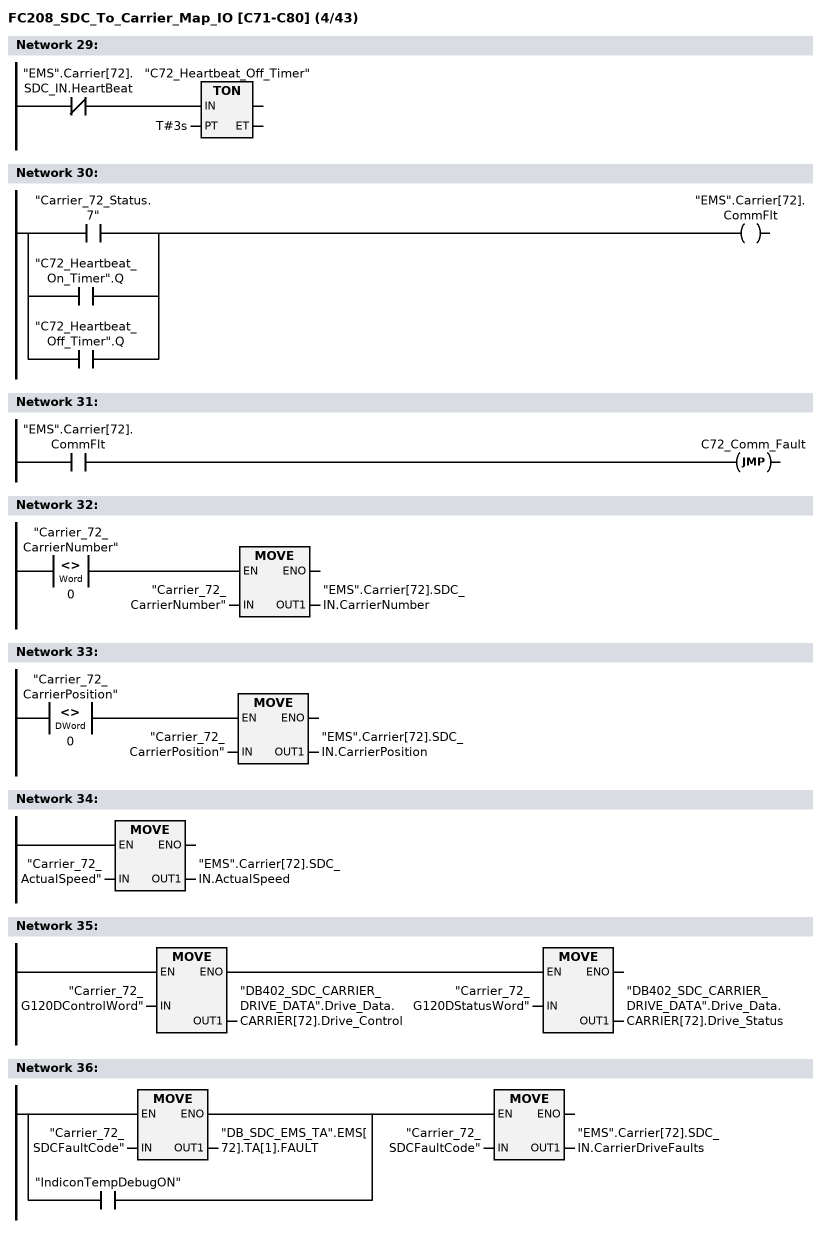
   "C72_Heartbeat_Off_Timer".TON(IN := NOT "EMS".Carrier[72].SDC_IN.HeartBeat, PT := T#3s);
END_REGION

REGION Network 30
   RUNG wire#powerrail
      Contact( "Carrier_72_Status.7" )
      wire#w1
      Coil( "EMS".Carrier[72].CommFlt )
   END_RUNG
   RUNG wire#powerrail
      Contact( "C72_Heartbeat_On_Timer".Q )
   END_RUNG wire#w1
   RUNG wire#powerrail
      Contact( "C72_Heartbeat_Off_Timer".Q )
   END_RUNG wire#w1
   // the same network as SCL:
   "EMS".Carrier[72].CommFlt := "Carrier_72_Status.7" OR "C72_Heartbeat_On_Timer".Q OR "C72_Heartbeat_Off_Timer".Q;
END_REGION

REGION Network 31
   RUNG wire#powerrail
      Contact( "EMS".Carrier[72].CommFlt )
      JumpCoil( C72_Comm_Fault )
   END_RUNG
   // the same network as SCL:
   IF "EMS".Carrier[72].CommFlt THEN GOTO C72_Comm_Fault; END_IF;
END_REGION

REGION Network 32
   RUNG wire#powerrail
      { S7_Templates := "SrcType := Word" } NE_Contact(in1 := "Carrier_72_CarrierNumber", in2 := 0)
      Move(in := "Carrier_72_CarrierNumber", out1 => "EMS".Carrier[72].SDC_IN.CarrierNumber)
   END_RUNG
   // the same network as SCL:
   IF "Carrier_72_CarrierNumber" <> 0 THEN
       "EMS".Carrier[72].SDC_IN.CarrierNumber := "Carrier_72_CarrierNumber";
   END_IF;
END_REGION

REGION Network 33
   RUNG wire#powerrail
      { S7_Templates := "SrcType := DWord" } NE_Contact(in1 := "Carrier_72_CarrierPosition", in2 := 0)
      Move(in := "Carrier_72_CarrierPosition", out1 => "EMS".Carrier[72].SDC_IN.CarrierPosition)
   END_RUNG
   // the same network as SCL:
   IF "Carrier_72_CarrierPosition" <> 0 THEN
       "EMS".Carrier[72].SDC_IN.CarrierPosition := "Carrier_72_CarrierPosition";
   END_IF;
END_REGION

REGION Network 34
   RUNG wire#powerrail
      Move(in := "Carrier_72_ActualSpeed", out1 => "EMS".Carrier[72].SDC_IN.ActualSpeed)
   END_RUNG
   // the same network as SCL:
   "EMS".Carrier[72].SDC_IN.ActualSpeed := "Carrier_72_ActualSpeed";
END_REGION

REGION Network 35
   RUNG wire#powerrail
      Move(in := "Carrier_72_G120DControlWord", out1 => "DB402_SDC_CARRIER_DRIVE_DATA".Drive_Data.CARRIER[72].Drive_Control)
      Move(in := "Carrier_72_G120DStatusWord", out1 => "DB402_SDC_CARRIER_DRIVE_DATA".Drive_Data.CARRIER[72].Drive_Status)
   END_RUNG
   // the same network as SCL:
   "DB402_SDC_CARRIER_DRIVE_DATA".Drive_Data.CARRIER[72].Drive_Control := "Carrier_72_G120DControlWord";
   "DB402_SDC_CARRIER_DRIVE_DATA".Drive_Data.CARRIER[72].Drive_Status := "Carrier_72_G120DStatusWord";
END_REGION

REGION Network 36
   RUNG wire#powerrail
      Move(in := "Carrier_72_SDCFaultCode", out1 => "DB_SDC_EMS_TA".EMS[72].TA[1].FAULT)
      wire#w1
      Move(in := "Carrier_72_SDCFaultCode", out1 => "EMS".Carrier[72].SDC_IN.CarrierDriveFaults)
   END_RUNG
   RUNG wire#powerrail
      Contact( "IndiconTempDebugON" )
   END_RUNG wire#w1
   // the same network as SCL:
   "DB_SDC_EMS_TA".EMS[72].TA[1].FAULT := "Carrier_72_SDCFaultCode";
   IF TRUE OR "IndiconTempDebugON" THEN
       "EMS".Carrier[72].SDC_IN.CarrierDriveFaults := "Carrier_72_SDCFaultCode";
   END_IF;
END_REGION

REGION Network 37
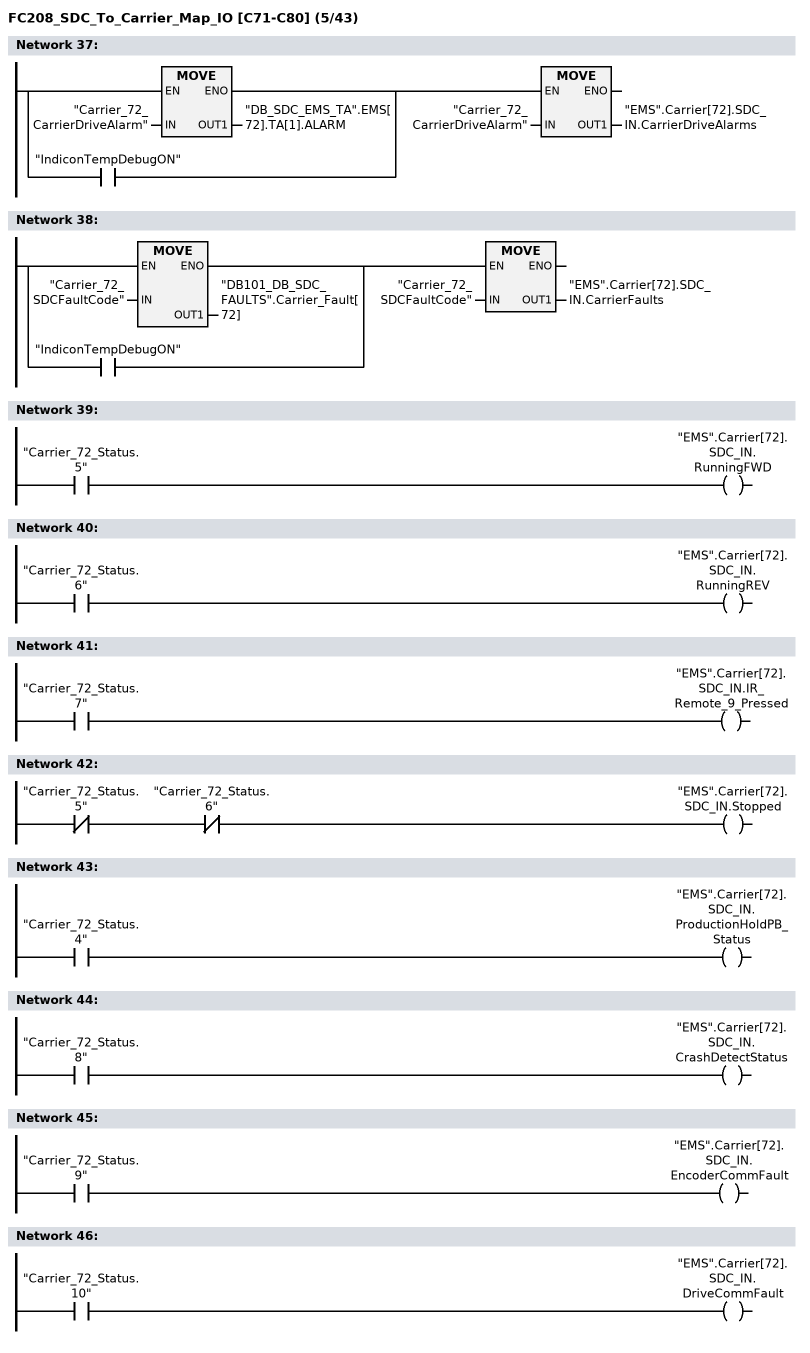
   RUNG wire#powerrail
      Move(in := "Carrier_72_CarrierDriveAlarm", out1 => "DB_SDC_EMS_TA".EMS[72].TA[1].ALARM)
      wire#w1
      Move(in := "Carrier_72_CarrierDriveAlarm", out1 => "EMS".Carrier[72].SDC_IN.CarrierDriveAlarms)
   END_RUNG
   RUNG wire#powerrail
      Contact( "IndiconTempDebugON" )
   END_RUNG wire#w1
   // the same network as SCL:
   "DB_SDC_EMS_TA".EMS[72].TA[1].ALARM := "Carrier_72_CarrierDriveAlarm";
   IF TRUE OR "IndiconTempDebugON" THEN
       "EMS".Carrier[72].SDC_IN.CarrierDriveAlarms := "Carrier_72_CarrierDriveAlarm";
   END_IF;
END_REGION

REGION Network 38
   RUNG wire#powerrail
      Move(in := "Carrier_72_SDCFaultCode", out1 => "DB101_DB_SDC_FAULTS".Carrier_Fault[72])
      wire#w1
      Move(in := "Carrier_72_SDCFaultCode", out1 => "EMS".Carrier[72].SDC_IN.CarrierFaults)
   END_RUNG
   RUNG wire#powerrail
      Contact( "IndiconTempDebugON" )
   END_RUNG wire#w1
   // the same network as SCL:
   "DB101_DB_SDC_FAULTS".Carrier_Fault[72] := "Carrier_72_SDCFaultCode";
   IF TRUE OR "IndiconTempDebugON" THEN
       "EMS".Carrier[72].SDC_IN.CarrierFaults := "Carrier_72_SDCFaultCode";
   END_IF;
END_REGION

REGION Network 39
   RUNG wire#powerrail
      Contact( "Carrier_72_Status.5" )
      Coil( "EMS".Carrier[72].SDC_IN.RunningFWD )
   END_RUNG
   // the same network as SCL:
   "EMS".Carrier[72].SDC_IN.RunningFWD := "Carrier_72_Status.5";
END_REGION

REGION Network 40
   RUNG wire#powerrail
      Contact( "Carrier_72_Status.6" )
      Coil( "EMS".Carrier[72].SDC_IN.RunningREV )
   END_RUNG
   // the same network as SCL:
   "EMS".Carrier[72].SDC_IN.RunningREV := "Carrier_72_Status.6";
END_REGION

REGION Network 41
   RUNG wire#powerrail
      Contact( "Carrier_72_Status.7" )
      Coil( "EMS".Carrier[72].SDC_IN.IR_Remote_9_Pressed )
   END_RUNG
   // the same network as SCL:
   "EMS".Carrier[72].SDC_IN.IR_Remote_9_Pressed := "Carrier_72_Status.7";
END_REGION

REGION Network 42
   RUNG wire#powerrail
      I_Contact( "Carrier_72_Status.5" )
      I_Contact( "Carrier_72_Status.6" )
      Coil( "EMS".Carrier[72].SDC_IN.Stopped )
   END_RUNG
   // the same network as SCL:
   "EMS".Carrier[72].SDC_IN.Stopped := NOT "Carrier_72_Status.5" AND NOT "Carrier_72_Status.6";
END_REGION

REGION Network 43
   RUNG wire#powerrail
      Contact( "Carrier_72_Status.4" )
      Coil( "EMS".Carrier[72].SDC_IN.ProductionHoldPB_Status )
   END_RUNG
   // the same network as SCL:
   "EMS".Carrier[72].SDC_IN.ProductionHoldPB_Status := "Carrier_72_Status.4";
END_REGION

REGION Network 44
   RUNG wire#powerrail
      Contact( "Carrier_72_Status.8" )
      Coil( "EMS".Carrier[72].SDC_IN.CrashDetectStatus )
   END_RUNG
   // the same network as SCL:
   "EMS".Carrier[72].SDC_IN.CrashDetectStatus := "Carrier_72_Status.8";
END_REGION

REGION Network 45
   RUNG wire#powerrail
      Contact( "Carrier_72_Status.9" )
      Coil( "EMS".Carrier[72].SDC_IN.EncoderCommFault )
   END_RUNG
   // the same network as SCL:
   "EMS".Carrier[72].SDC_IN.EncoderCommFault := "Carrier_72_Status.9";
END_REGION

REGION Network 46
   RUNG wire#powerrail
      Contact( "Carrier_72_Status.10" )
      Coil( "EMS".Carrier[72].SDC_IN.DriveCommFault )
   END_RUNG
   // the same network as SCL:
   "EMS".Carrier[72].SDC_IN.DriveCommFault := "Carrier_72_Status.10";
END_REGION

REGION Network 47
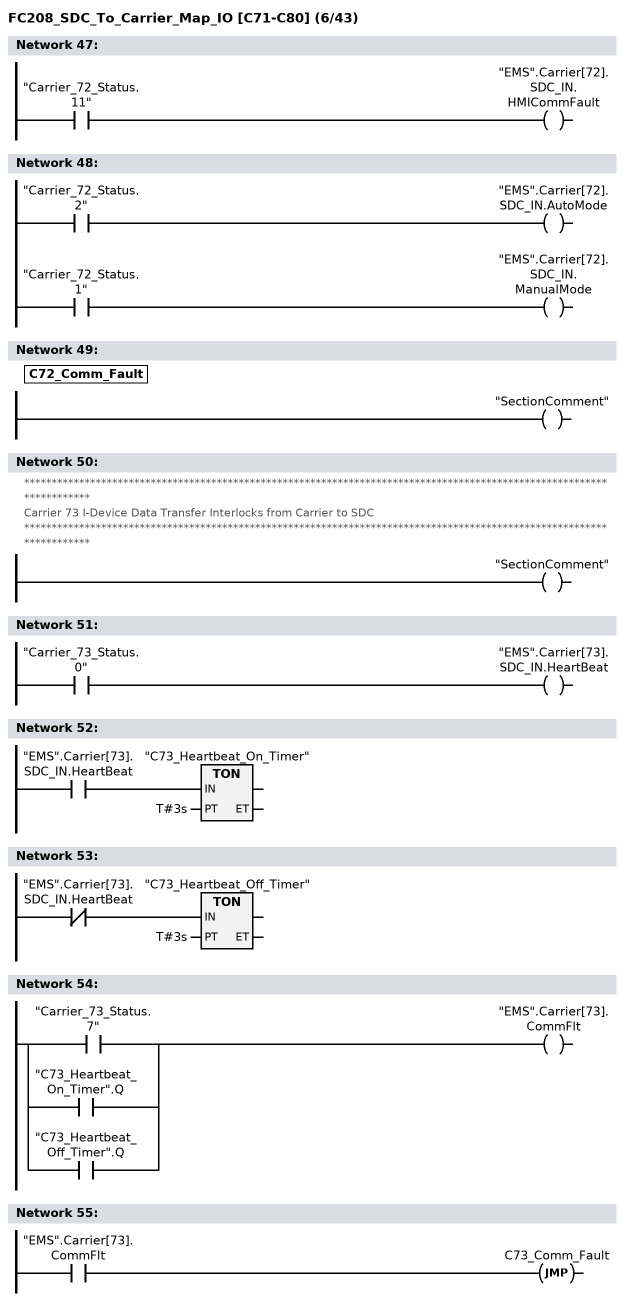
   RUNG wire#powerrail
      Contact( "Carrier_72_Status.11" )
      Coil( "EMS".Carrier[72].SDC_IN.HMICommFault )
   END_RUNG
   // the same network as SCL:
   "EMS".Carrier[72].SDC_IN.HMICommFault := "Carrier_72_Status.11";
END_REGION

REGION Network 48
   RUNG wire#powerrail
      Contact( "Carrier_72_Status.2" )
      Coil( "EMS".Carrier[72].SDC_IN.AutoMode )
   END_RUNG
   RUNG wire#powerrail
      Contact( "Carrier_72_Status.1" )
      Coil( "EMS".Carrier[72].SDC_IN.ManualMode )
   END_RUNG
   // the same network as SCL:
   "EMS".Carrier[72].SDC_IN.AutoMode := "Carrier_72_Status.2";
   "EMS".Carrier[72].SDC_IN.ManualMode := "Carrier_72_Status.1";
END_REGION

REGION Network 49
   Label( C72_Comm_Fault )
   RUNG wire#powerrail
      Coil( "SectionComment" )
   END_RUNG
   // the same network as SCL:
   C72_Comm_Fault:
   "SectionComment" := TRUE;
END_REGION

REGION Network 50
   // **********************************************************************************************************************
   // 
   // Carrier 73 I-Device Data Transfer Interlocks from Carrier to SDC
   // 
   // **********************************************************************************************************************
   RUNG wire#powerrail
      Coil( "SectionComment" )
   END_RUNG
   // the same network as SCL:
   "SectionComment" := TRUE;
END_REGION

REGION Network 51
   RUNG wire#powerrail
      Contact( "Carrier_73_Status.0" )
      Coil( "EMS".Carrier[73].SDC_IN.HeartBeat )
   END_RUNG
   // the same network as SCL:
   "EMS".Carrier[73].SDC_IN.HeartBeat := "Carrier_73_Status.0";
END_REGION

REGION Network 52
   "C73_Heartbeat_On_Timer".TON(IN := "EMS".Carrier[73].SDC_IN.HeartBeat, PT := T#3s);
END_REGION

REGION Network 53
   "C73_Heartbeat_Off_Timer".TON(IN := NOT "EMS".Carrier[73].SDC_IN.HeartBeat, PT := T#3s);
END_REGION

REGION Network 54
   RUNG wire#powerrail
      Contact( "Carrier_73_Status.7" )
      wire#w1
      Coil( "EMS".Carrier[73].CommFlt )
   END_RUNG
   RUNG wire#powerrail
      Contact( "C73_Heartbeat_On_Timer".Q )
   END_RUNG wire#w1
   RUNG wire#powerrail
      Contact( "C73_Heartbeat_Off_Timer".Q )
   END_RUNG wire#w1
   // the same network as SCL:
   "EMS".Carrier[73].CommFlt := "Carrier_73_Status.7" OR "C73_Heartbeat_On_Timer".Q OR "C73_Heartbeat_Off_Timer".Q;
END_REGION

REGION Network 55
   RUNG wire#powerrail
      Contact( "EMS".Carrier[73].CommFlt )
      JumpCoil( C73_Comm_Fault )
   END_RUNG
   // the same network as SCL:
   IF "EMS".Carrier[73].CommFlt THEN GOTO C73_Comm_Fault; END_IF;
END_REGION

REGION Network 56
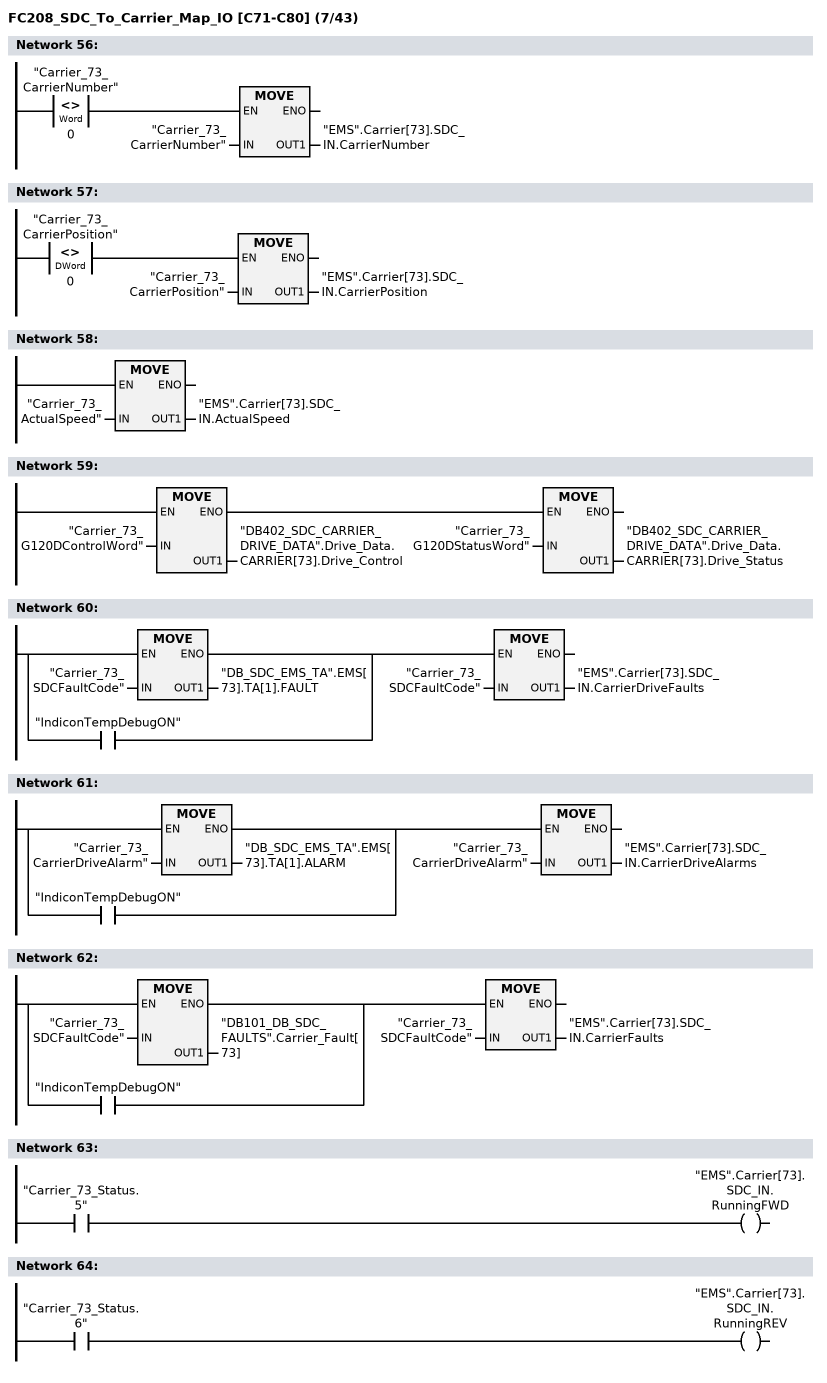
   RUNG wire#powerrail
      { S7_Templates := "SrcType := Word" } NE_Contact(in1 := "Carrier_73_CarrierNumber", in2 := 0)
      Move(in := "Carrier_73_CarrierNumber", out1 => "EMS".Carrier[73].SDC_IN.CarrierNumber)
   END_RUNG
   // the same network as SCL:
   IF "Carrier_73_CarrierNumber" <> 0 THEN
       "EMS".Carrier[73].SDC_IN.CarrierNumber := "Carrier_73_CarrierNumber";
   END_IF;
END_REGION

REGION Network 57
   RUNG wire#powerrail
      { S7_Templates := "SrcType := DWord" } NE_Contact(in1 := "Carrier_73_CarrierPosition", in2 := 0)
      Move(in := "Carrier_73_CarrierPosition", out1 => "EMS".Carrier[73].SDC_IN.CarrierPosition)
   END_RUNG
   // the same network as SCL:
   IF "Carrier_73_CarrierPosition" <> 0 THEN
       "EMS".Carrier[73].SDC_IN.CarrierPosition := "Carrier_73_CarrierPosition";
   END_IF;
END_REGION

REGION Network 58
   RUNG wire#powerrail
      Move(in := "Carrier_73_ActualSpeed", out1 => "EMS".Carrier[73].SDC_IN.ActualSpeed)
   END_RUNG
   // the same network as SCL:
   "EMS".Carrier[73].SDC_IN.ActualSpeed := "Carrier_73_ActualSpeed";
END_REGION

REGION Network 59
   RUNG wire#powerrail
      Move(in := "Carrier_73_G120DControlWord", out1 => "DB402_SDC_CARRIER_DRIVE_DATA".Drive_Data.CARRIER[73].Drive_Control)
      Move(in := "Carrier_73_G120DStatusWord", out1 => "DB402_SDC_CARRIER_DRIVE_DATA".Drive_Data.CARRIER[73].Drive_Status)
   END_RUNG
   // the same network as SCL:
   "DB402_SDC_CARRIER_DRIVE_DATA".Drive_Data.CARRIER[73].Drive_Control := "Carrier_73_G120DControlWord";
   "DB402_SDC_CARRIER_DRIVE_DATA".Drive_Data.CARRIER[73].Drive_Status := "Carrier_73_G120DStatusWord";
END_REGION

REGION Network 60
   RUNG wire#powerrail
      Move(in := "Carrier_73_SDCFaultCode", out1 => "DB_SDC_EMS_TA".EMS[73].TA[1].FAULT)
      wire#w1
      Move(in := "Carrier_73_SDCFaultCode", out1 => "EMS".Carrier[73].SDC_IN.CarrierDriveFaults)
   END_RUNG
   RUNG wire#powerrail
      Contact( "IndiconTempDebugON" )
   END_RUNG wire#w1
   // the same network as SCL:
   "DB_SDC_EMS_TA".EMS[73].TA[1].FAULT := "Carrier_73_SDCFaultCode";
   IF TRUE OR "IndiconTempDebugON" THEN
       "EMS".Carrier[73].SDC_IN.CarrierDriveFaults := "Carrier_73_SDCFaultCode";
   END_IF;
END_REGION

REGION Network 61
   RUNG wire#powerrail
      Move(in := "Carrier_73_CarrierDriveAlarm", out1 => "DB_SDC_EMS_TA".EMS[73].TA[1].ALARM)
      wire#w1
      Move(in := "Carrier_73_CarrierDriveAlarm", out1 => "EMS".Carrier[73].SDC_IN.CarrierDriveAlarms)
   END_RUNG
   RUNG wire#powerrail
      Contact( "IndiconTempDebugON" )
   END_RUNG wire#w1
   // the same network as SCL:
   "DB_SDC_EMS_TA".EMS[73].TA[1].ALARM := "Carrier_73_CarrierDriveAlarm";
   IF TRUE OR "IndiconTempDebugON" THEN
       "EMS".Carrier[73].SDC_IN.CarrierDriveAlarms := "Carrier_73_CarrierDriveAlarm";
   END_IF;
END_REGION

REGION Network 62
   RUNG wire#powerrail
      Move(in := "Carrier_73_SDCFaultCode", out1 => "DB101_DB_SDC_FAULTS".Carrier_Fault[73])
      wire#w1
      Move(in := "Carrier_73_SDCFaultCode", out1 => "EMS".Carrier[73].SDC_IN.CarrierFaults)
   END_RUNG
   RUNG wire#powerrail
      Contact( "IndiconTempDebugON" )
   END_RUNG wire#w1
   // the same network as SCL:
   "DB101_DB_SDC_FAULTS".Carrier_Fault[73] := "Carrier_73_SDCFaultCode";
   IF TRUE OR "IndiconTempDebugON" THEN
       "EMS".Carrier[73].SDC_IN.CarrierFaults := "Carrier_73_SDCFaultCode";
   END_IF;
END_REGION

REGION Network 63
   RUNG wire#powerrail
      Contact( "Carrier_73_Status.5" )
      Coil( "EMS".Carrier[73].SDC_IN.RunningFWD )
   END_RUNG
   // the same network as SCL:
   "EMS".Carrier[73].SDC_IN.RunningFWD := "Carrier_73_Status.5";
END_REGION

REGION Network 64
   RUNG wire#powerrail
      Contact( "Carrier_73_Status.6" )
      Coil( "EMS".Carrier[73].SDC_IN.RunningREV )
   END_RUNG
   // the same network as SCL:
   "EMS".Carrier[73].SDC_IN.RunningREV := "Carrier_73_Status.6";
END_REGION

REGION Network 65
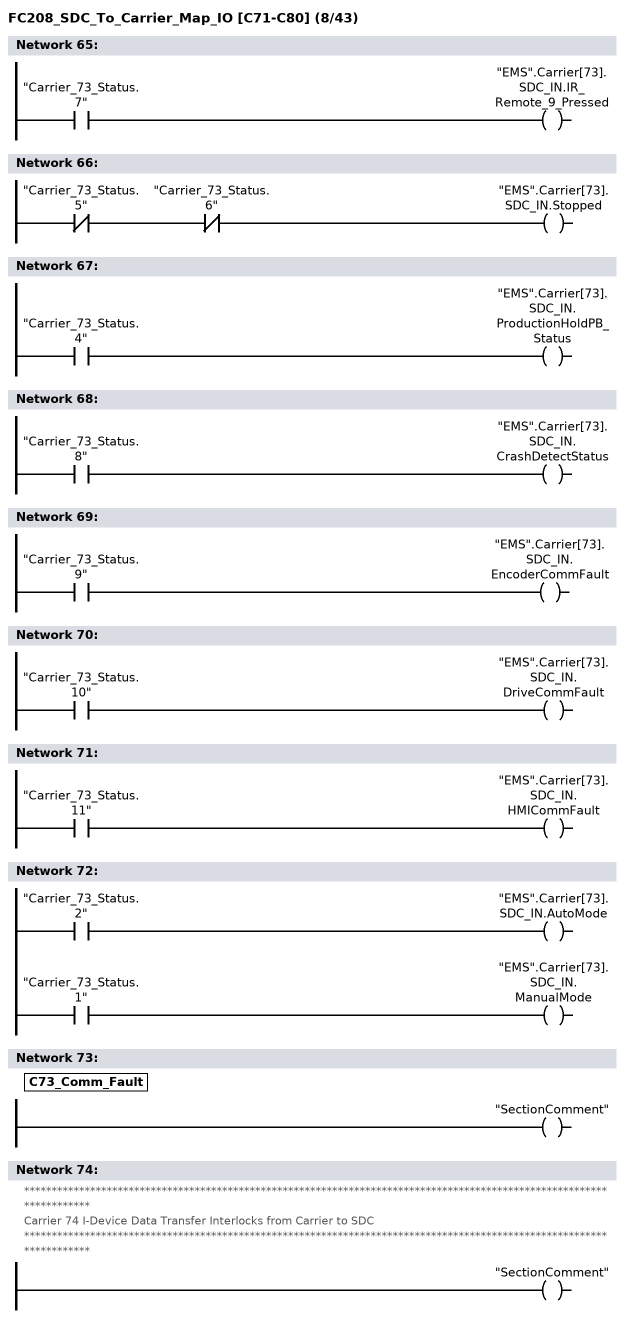
   RUNG wire#powerrail
      Contact( "Carrier_73_Status.7" )
      Coil( "EMS".Carrier[73].SDC_IN.IR_Remote_9_Pressed )
   END_RUNG
   // the same network as SCL:
   "EMS".Carrier[73].SDC_IN.IR_Remote_9_Pressed := "Carrier_73_Status.7";
END_REGION

REGION Network 66
   RUNG wire#powerrail
      I_Contact( "Carrier_73_Status.5" )
      I_Contact( "Carrier_73_Status.6" )
      Coil( "EMS".Carrier[73].SDC_IN.Stopped )
   END_RUNG
   // the same network as SCL:
   "EMS".Carrier[73].SDC_IN.Stopped := NOT "Carrier_73_Status.5" AND NOT "Carrier_73_Status.6";
END_REGION

REGION Network 67
   RUNG wire#powerrail
      Contact( "Carrier_73_Status.4" )
      Coil( "EMS".Carrier[73].SDC_IN.ProductionHoldPB_Status )
   END_RUNG
   // the same network as SCL:
   "EMS".Carrier[73].SDC_IN.ProductionHoldPB_Status := "Carrier_73_Status.4";
END_REGION

REGION Network 68
   RUNG wire#powerrail
      Contact( "Carrier_73_Status.8" )
      Coil( "EMS".Carrier[73].SDC_IN.CrashDetectStatus )
   END_RUNG
   // the same network as SCL:
   "EMS".Carrier[73].SDC_IN.CrashDetectStatus := "Carrier_73_Status.8";
END_REGION

REGION Network 69
   RUNG wire#powerrail
      Contact( "Carrier_73_Status.9" )
      Coil( "EMS".Carrier[73].SDC_IN.EncoderCommFault )
   END_RUNG
   // the same network as SCL:
   "EMS".Carrier[73].SDC_IN.EncoderCommFault := "Carrier_73_Status.9";
END_REGION

REGION Network 70
   RUNG wire#powerrail
      Contact( "Carrier_73_Status.10" )
      Coil( "EMS".Carrier[73].SDC_IN.DriveCommFault )
   END_RUNG
   // the same network as SCL:
   "EMS".Carrier[73].SDC_IN.DriveCommFault := "Carrier_73_Status.10";
END_REGION

REGION Network 71
   RUNG wire#powerrail
      Contact( "Carrier_73_Status.11" )
      Coil( "EMS".Carrier[73].SDC_IN.HMICommFault )
   END_RUNG
   // the same network as SCL:
   "EMS".Carrier[73].SDC_IN.HMICommFault := "Carrier_73_Status.11";
END_REGION

REGION Network 72
   RUNG wire#powerrail
      Contact( "Carrier_73_Status.2" )
      Coil( "EMS".Carrier[73].SDC_IN.AutoMode )
   END_RUNG
   RUNG wire#powerrail
      Contact( "Carrier_73_Status.1" )
      Coil( "EMS".Carrier[73].SDC_IN.ManualMode )
   END_RUNG
   // the same network as SCL:
   "EMS".Carrier[73].SDC_IN.AutoMode := "Carrier_73_Status.2";
   "EMS".Carrier[73].SDC_IN.ManualMode := "Carrier_73_Status.1";
END_REGION

REGION Network 73
   Label( C73_Comm_Fault )
   RUNG wire#powerrail
      Coil( "SectionComment" )
   END_RUNG
   // the same network as SCL:
   C73_Comm_Fault:
   "SectionComment" := TRUE;
END_REGION

REGION Network 74
   // **********************************************************************************************************************
   // 
   // Carrier 74 I-Device Data Transfer Interlocks from Carrier to SDC
   // 
   // **********************************************************************************************************************
   RUNG wire#powerrail
      Coil( "SectionComment" )
   END_RUNG
   // the same network as SCL:
   "SectionComment" := TRUE;
END_REGION

REGION Network 75
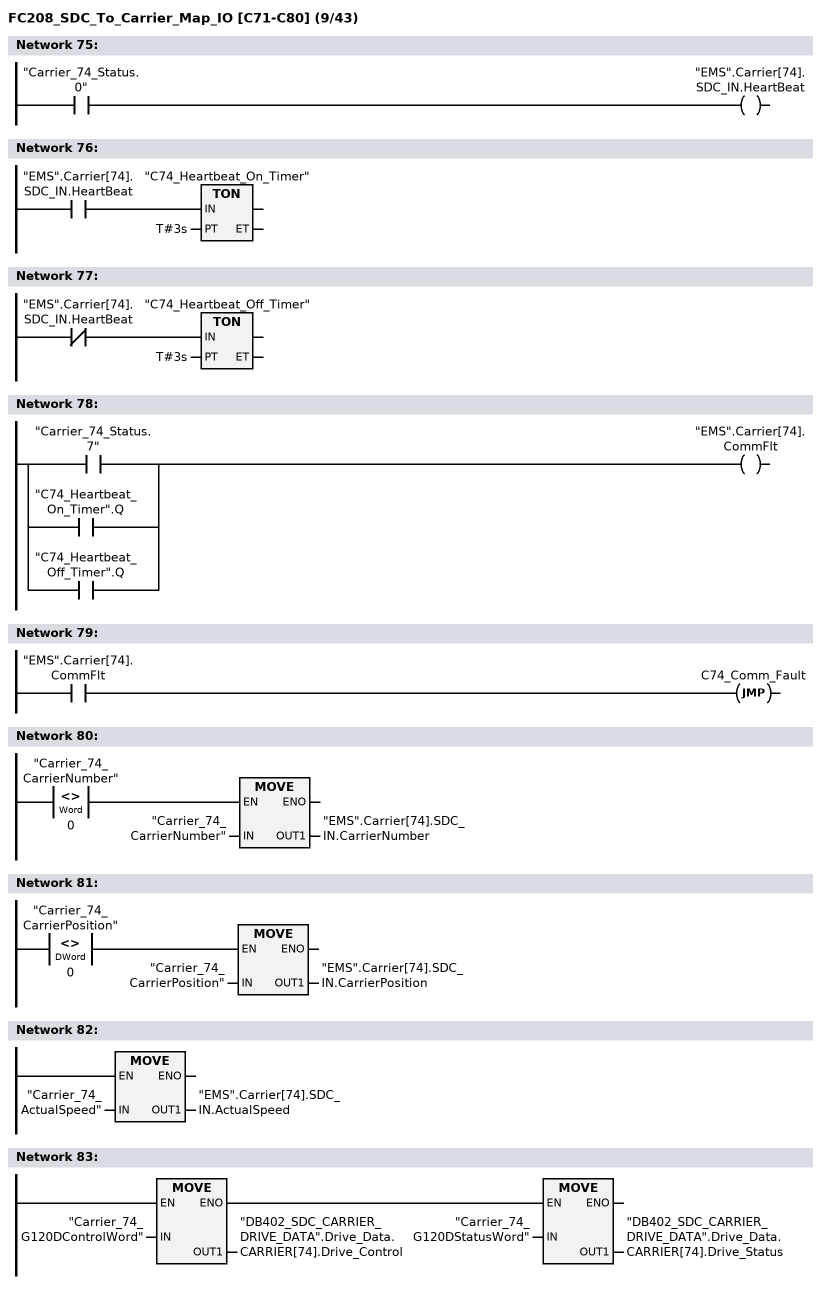
   RUNG wire#powerrail
      Contact( "Carrier_74_Status.0" )
      Coil( "EMS".Carrier[74].SDC_IN.HeartBeat )
   END_RUNG
   // the same network as SCL:
   "EMS".Carrier[74].SDC_IN.HeartBeat := "Carrier_74_Status.0";
END_REGION

REGION Network 76
   "C74_Heartbeat_On_Timer".TON(IN := "EMS".Carrier[74].SDC_IN.HeartBeat, PT := T#3s);
END_REGION

REGION Network 77
   "C74_Heartbeat_Off_Timer".TON(IN := NOT "EMS".Carrier[74].SDC_IN.HeartBeat, PT := T#3s);
END_REGION

REGION Network 78
   RUNG wire#powerrail
      Contact( "Carrier_74_Status.7" )
      wire#w1
      Coil( "EMS".Carrier[74].CommFlt )
   END_RUNG
   RUNG wire#powerrail
      Contact( "C74_Heartbeat_On_Timer".Q )
   END_RUNG wire#w1
   RUNG wire#powerrail
      Contact( "C74_Heartbeat_Off_Timer".Q )
   END_RUNG wire#w1
   // the same network as SCL:
   "EMS".Carrier[74].CommFlt := "Carrier_74_Status.7" OR "C74_Heartbeat_On_Timer".Q OR "C74_Heartbeat_Off_Timer".Q;
END_REGION

REGION Network 79
   RUNG wire#powerrail
      Contact( "EMS".Carrier[74].CommFlt )
      JumpCoil( C74_Comm_Fault )
   END_RUNG
   // the same network as SCL:
   IF "EMS".Carrier[74].CommFlt THEN GOTO C74_Comm_Fault; END_IF;
END_REGION

REGION Network 80
   RUNG wire#powerrail
      { S7_Templates := "SrcType := Word" } NE_Contact(in1 := "Carrier_74_CarrierNumber", in2 := 0)
      Move(in := "Carrier_74_CarrierNumber", out1 => "EMS".Carrier[74].SDC_IN.CarrierNumber)
   END_RUNG
   // the same network as SCL:
   IF "Carrier_74_CarrierNumber" <> 0 THEN
       "EMS".Carrier[74].SDC_IN.CarrierNumber := "Carrier_74_CarrierNumber";
   END_IF;
END_REGION

REGION Network 81
   RUNG wire#powerrail
      { S7_Templates := "SrcType := DWord" } NE_Contact(in1 := "Carrier_74_CarrierPosition", in2 := 0)
      Move(in := "Carrier_74_CarrierPosition", out1 => "EMS".Carrier[74].SDC_IN.CarrierPosition)
   END_RUNG
   // the same network as SCL:
   IF "Carrier_74_CarrierPosition" <> 0 THEN
       "EMS".Carrier[74].SDC_IN.CarrierPosition := "Carrier_74_CarrierPosition";
   END_IF;
END_REGION

REGION Network 82
   RUNG wire#powerrail
      Move(in := "Carrier_74_ActualSpeed", out1 => "EMS".Carrier[74].SDC_IN.ActualSpeed)
   END_RUNG
   // the same network as SCL:
   "EMS".Carrier[74].SDC_IN.ActualSpeed := "Carrier_74_ActualSpeed";
END_REGION

REGION Network 83
   RUNG wire#powerrail
      Move(in := "Carrier_74_G120DControlWord", out1 => "DB402_SDC_CARRIER_DRIVE_DATA".Drive_Data.CARRIER[74].Drive_Control)
      Move(in := "Carrier_74_G120DStatusWord", out1 => "DB402_SDC_CARRIER_DRIVE_DATA".Drive_Data.CARRIER[74].Drive_Status)
   END_RUNG
   // the same network as SCL:
   "DB402_SDC_CARRIER_DRIVE_DATA".Drive_Data.CARRIER[74].Drive_Control := "Carrier_74_G120DControlWord";
   "DB402_SDC_CARRIER_DRIVE_DATA".Drive_Data.CARRIER[74].Drive_Status := "Carrier_74_G120DStatusWord";
END_REGION

REGION Network 84
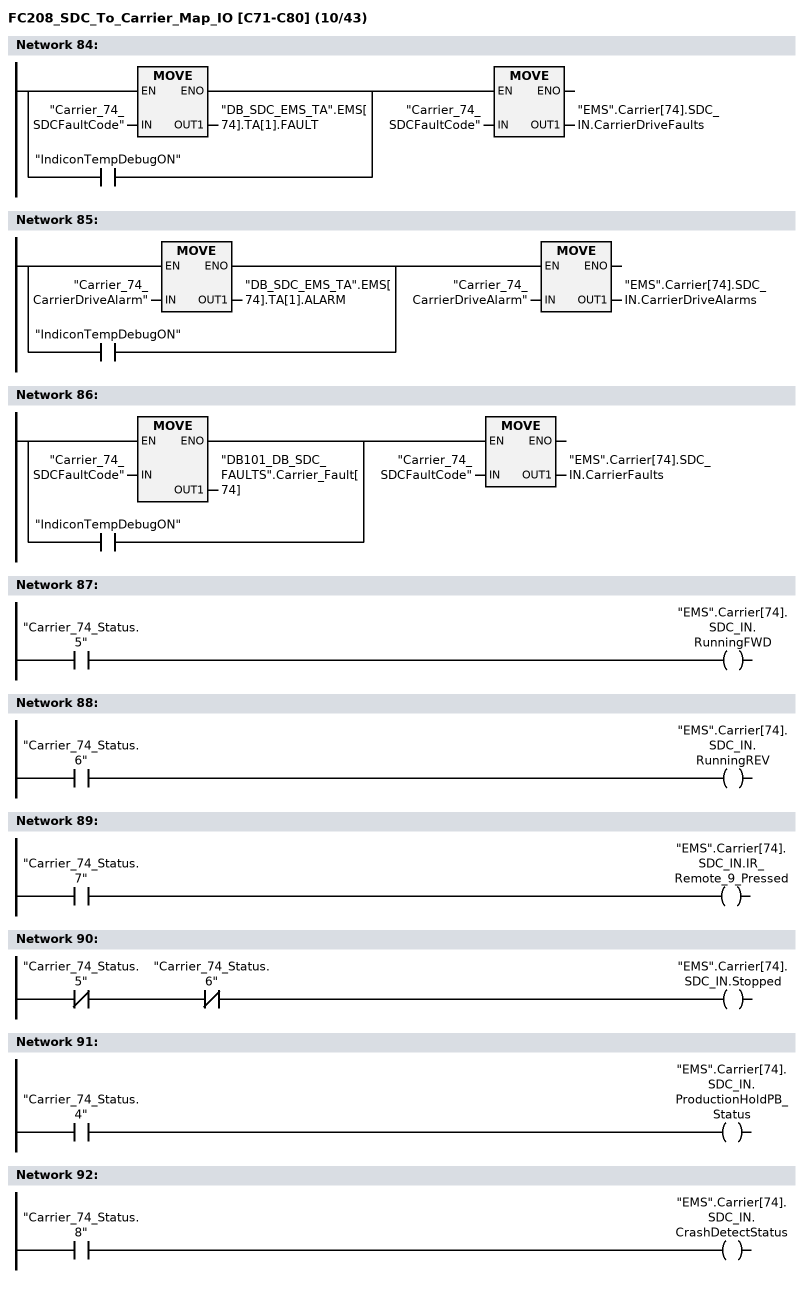
   RUNG wire#powerrail
      Move(in := "Carrier_74_SDCFaultCode", out1 => "DB_SDC_EMS_TA".EMS[74].TA[1].FAULT)
      wire#w1
      Move(in := "Carrier_74_SDCFaultCode", out1 => "EMS".Carrier[74].SDC_IN.CarrierDriveFaults)
   END_RUNG
   RUNG wire#powerrail
      Contact( "IndiconTempDebugON" )
   END_RUNG wire#w1
   // the same network as SCL:
   "DB_SDC_EMS_TA".EMS[74].TA[1].FAULT := "Carrier_74_SDCFaultCode";
   IF TRUE OR "IndiconTempDebugON" THEN
       "EMS".Carrier[74].SDC_IN.CarrierDriveFaults := "Carrier_74_SDCFaultCode";
   END_IF;
END_REGION

REGION Network 85
   RUNG wire#powerrail
      Move(in := "Carrier_74_CarrierDriveAlarm", out1 => "DB_SDC_EMS_TA".EMS[74].TA[1].ALARM)
      wire#w1
      Move(in := "Carrier_74_CarrierDriveAlarm", out1 => "EMS".Carrier[74].SDC_IN.CarrierDriveAlarms)
   END_RUNG
   RUNG wire#powerrail
      Contact( "IndiconTempDebugON" )
   END_RUNG wire#w1
   // the same network as SCL:
   "DB_SDC_EMS_TA".EMS[74].TA[1].ALARM := "Carrier_74_CarrierDriveAlarm";
   IF TRUE OR "IndiconTempDebugON" THEN
       "EMS".Carrier[74].SDC_IN.CarrierDriveAlarms := "Carrier_74_CarrierDriveAlarm";
   END_IF;
END_REGION

REGION Network 86
   RUNG wire#powerrail
      Move(in := "Carrier_74_SDCFaultCode", out1 => "DB101_DB_SDC_FAULTS".Carrier_Fault[74])
      wire#w1
      Move(in := "Carrier_74_SDCFaultCode", out1 => "EMS".Carrier[74].SDC_IN.CarrierFaults)
   END_RUNG
   RUNG wire#powerrail
      Contact( "IndiconTempDebugON" )
   END_RUNG wire#w1
   // the same network as SCL:
   "DB101_DB_SDC_FAULTS".Carrier_Fault[74] := "Carrier_74_SDCFaultCode";
   IF TRUE OR "IndiconTempDebugON" THEN
       "EMS".Carrier[74].SDC_IN.CarrierFaults := "Carrier_74_SDCFaultCode";
   END_IF;
END_REGION

REGION Network 87
   RUNG wire#powerrail
      Contact( "Carrier_74_Status.5" )
      Coil( "EMS".Carrier[74].SDC_IN.RunningFWD )
   END_RUNG
   // the same network as SCL:
   "EMS".Carrier[74].SDC_IN.RunningFWD := "Carrier_74_Status.5";
END_REGION

REGION Network 88
   RUNG wire#powerrail
      Contact( "Carrier_74_Status.6" )
      Coil( "EMS".Carrier[74].SDC_IN.RunningREV )
   END_RUNG
   // the same network as SCL:
   "EMS".Carrier[74].SDC_IN.RunningREV := "Carrier_74_Status.6";
END_REGION

REGION Network 89
   RUNG wire#powerrail
      Contact( "Carrier_74_Status.7" )
      Coil( "EMS".Carrier[74].SDC_IN.IR_Remote_9_Pressed )
   END_RUNG
   // the same network as SCL:
   "EMS".Carrier[74].SDC_IN.IR_Remote_9_Pressed := "Carrier_74_Status.7";
END_REGION

REGION Network 90
   RUNG wire#powerrail
      I_Contact( "Carrier_74_Status.5" )
      I_Contact( "Carrier_74_Status.6" )
      Coil( "EMS".Carrier[74].SDC_IN.Stopped )
   END_RUNG
   // the same network as SCL:
   "EMS".Carrier[74].SDC_IN.Stopped := NOT "Carrier_74_Status.5" AND NOT "Carrier_74_Status.6";
END_REGION

REGION Network 91
   RUNG wire#powerrail
      Contact( "Carrier_74_Status.4" )
      Coil( "EMS".Carrier[74].SDC_IN.ProductionHoldPB_Status )
   END_RUNG
   // the same network as SCL:
   "EMS".Carrier[74].SDC_IN.ProductionHoldPB_Status := "Carrier_74_Status.4";
END_REGION

REGION Network 92
   RUNG wire#powerrail
      Contact( "Carrier_74_Status.8" )
      Coil( "EMS".Carrier[74].SDC_IN.CrashDetectStatus )
   END_RUNG
   // the same network as SCL:
   "EMS".Carrier[74].SDC_IN.CrashDetectStatus := "Carrier_74_Status.8";
END_REGION

REGION Network 93
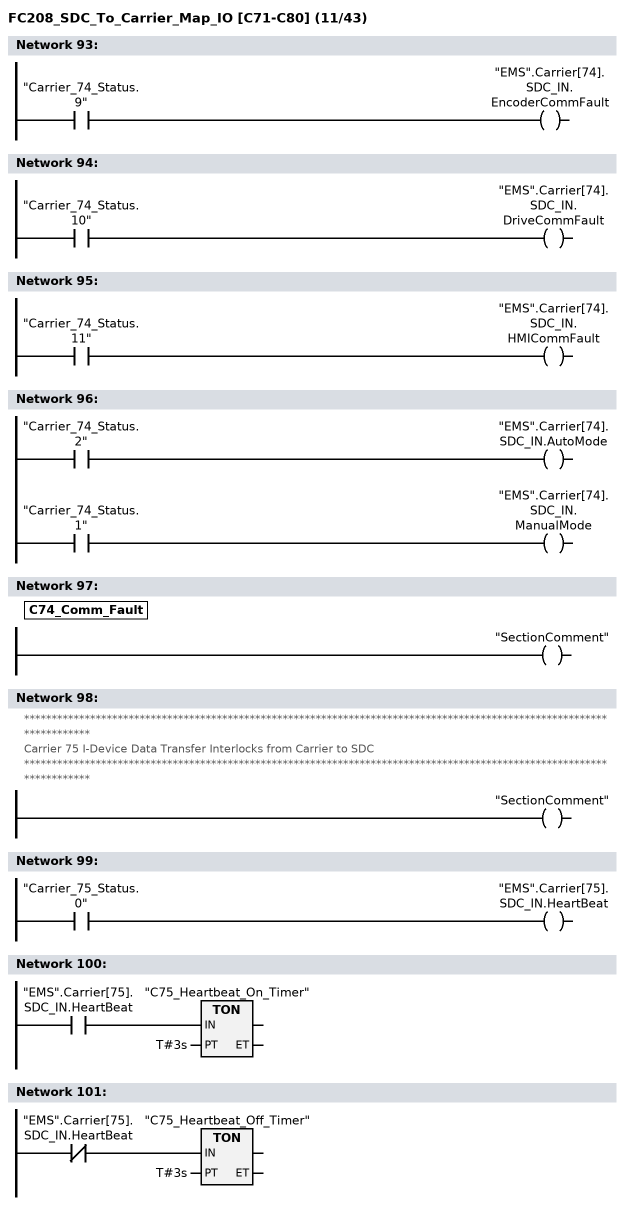
   RUNG wire#powerrail
      Contact( "Carrier_74_Status.9" )
      Coil( "EMS".Carrier[74].SDC_IN.EncoderCommFault )
   END_RUNG
   // the same network as SCL:
   "EMS".Carrier[74].SDC_IN.EncoderCommFault := "Carrier_74_Status.9";
END_REGION

REGION Network 94
   RUNG wire#powerrail
      Contact( "Carrier_74_Status.10" )
      Coil( "EMS".Carrier[74].SDC_IN.DriveCommFault )
   END_RUNG
   // the same network as SCL:
   "EMS".Carrier[74].SDC_IN.DriveCommFault := "Carrier_74_Status.10";
END_REGION

REGION Network 95
   RUNG wire#powerrail
      Contact( "Carrier_74_Status.11" )
      Coil( "EMS".Carrier[74].SDC_IN.HMICommFault )
   END_RUNG
   // the same network as SCL:
   "EMS".Carrier[74].SDC_IN.HMICommFault := "Carrier_74_Status.11";
END_REGION

REGION Network 96
   RUNG wire#powerrail
      Contact( "Carrier_74_Status.2" )
      Coil( "EMS".Carrier[74].SDC_IN.AutoMode )
   END_RUNG
   RUNG wire#powerrail
      Contact( "Carrier_74_Status.1" )
      Coil( "EMS".Carrier[74].SDC_IN.ManualMode )
   END_RUNG
   // the same network as SCL:
   "EMS".Carrier[74].SDC_IN.AutoMode := "Carrier_74_Status.2";
   "EMS".Carrier[74].SDC_IN.ManualMode := "Carrier_74_Status.1";
END_REGION

REGION Network 97
   Label( C74_Comm_Fault )
   RUNG wire#powerrail
      Coil( "SectionComment" )
   END_RUNG
   // the same network as SCL:
   C74_Comm_Fault:
   "SectionComment" := TRUE;
END_REGION

REGION Network 98
   // **********************************************************************************************************************
   // 
   // Carrier 75 I-Device Data Transfer Interlocks from Carrier to SDC
   // 
   // **********************************************************************************************************************
   RUNG wire#powerrail
      Coil( "SectionComment" )
   END_RUNG
   // the same network as SCL:
   "SectionComment" := TRUE;
END_REGION

REGION Network 99
   RUNG wire#powerrail
      Contact( "Carrier_75_Status.0" )
      Coil( "EMS".Carrier[75].SDC_IN.HeartBeat )
   END_RUNG
   // the same network as SCL:
   "EMS".Carrier[75].SDC_IN.HeartBeat := "Carrier_75_Status.0";
END_REGION

REGION Network 100
   "C75_Heartbeat_On_Timer".TON(IN := "EMS".Carrier[75].SDC_IN.HeartBeat, PT := T#3s);
END_REGION

REGION Network 101
   "C75_Heartbeat_Off_Timer".TON(IN := NOT "EMS".Carrier[75].SDC_IN.HeartBeat, PT := T#3s);
END_REGION

REGION Network 102
